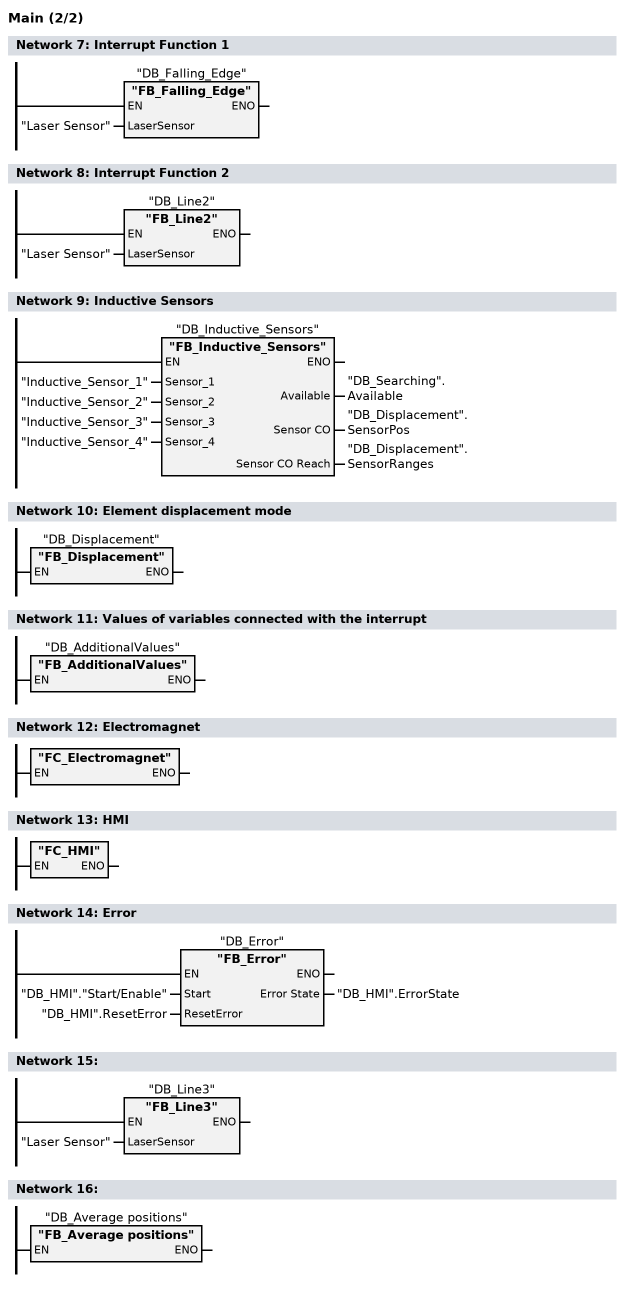
   RUNG wire#powerrail
      "DB_Falling_Edge"(LaserSensor := "Laser Sensor")
   END_RUNG
   // the same network as SCL:
   "DB_Falling_Edge"(LaserSensor := "Laser Sensor");   // "FB_Falling_Edge"
END_REGION

REGION Network 8: Interrupt Function 2
   RUNG wire#powerrail
      "DB_Line2"(LaserSensor := "Laser Sensor")
   END_RUNG
   // the same network as SCL:
   "DB_Line2"(LaserSensor := "Laser Sensor");   // "FB_Line2"
END_REGION

REGION Network 9: Inductive Sensors
   RUNG wire#powerrail
      "DB_Inductive_Sensors"(Sensor_1 := "Inductive_Sensor_1", Sensor_2 := "Inductive_Sensor_2", Sensor_3 := "Inductive_Sensor_3", Sensor_4 := "Inductive_Sensor_4", Available => "DB_Searching".Available, "Sensor CO" => "DB_Displacement".SensorPos, "Sensor CO Reach" => "DB_Displacement".SensorRanges)
   END_RUNG
   // the same network as SCL:
   "DB_Inductive_Sensors"(Sensor_1 := "Inductive_Sensor_1",   // "FB_Inductive_Sensors"
                          Sensor_2 := "Inductive_Sensor_2",
                          Sensor_3 := "Inductive_Sensor_3",
                          Sensor_4 := "Inductive_Sensor_4",
                          Available => "DB_Searching".Available,
                          "Sensor CO" => "DB_Displacement".SensorPos,
                          "Sensor CO Reach" => "DB_Displacement".SensorRanges);
END_REGION

REGION Network 10: Element displacement mode
   RUNG wire#powerrail
      "DB_Displacement"()
   END_RUNG
   // the same network as SCL:
   "DB_Displacement"();   // "FB_Displacement"
END_REGION

REGION Network 11: Values of variables connected with the interrupt
   RUNG wire#powerrail
      "DB_AdditionalValues"()
   END_RUNG
   // the same network as SCL:
   "DB_AdditionalValues"();   // "FB_AdditionalValues"
END_REGION

REGION Network 12: Electromagnet
   RUNG wire#powerrail
      "FC_Electromagnet"()
   END_RUNG
   // the same network as SCL:
   "FC_Electromagnet"();
END_REGION

REGION Network 13: HMI
   RUNG wire#powerrail
      "FC_HMI"()
   END_RUNG
   // the same network as SCL:
   "FC_HMI"();
END_REGION

REGION Network 14: Error
   RUNG wire#powerrail
      "DB_Error"(Start := "DB_HMI"."Start/Enable", ResetError := "DB_HMI".ResetError, "Error State" => "DB_HMI".ErrorState)
   END_RUNG
   // the same network as SCL:
   "DB_Error"(Start := "DB_HMI"."Start/Enable",   // "FB_Error"
              ResetError := "DB_HMI".ResetError,
              "Error State" => "DB_HMI".ErrorState);
END_REGION

REGION Network 15
   RUNG wire#powerrail
      "DB_Line3"(LaserSensor := "Laser Sensor")
   END_RUNG
   // the same network as SCL:
   "DB_Line3"(LaserSensor := "Laser Sensor");   // "FB_Line3"
END_REGION

REGION Network 16
   RUNG wire#powerrail
      "DB_Average positions"()
   END_RUNG
   // the same network as SCL:
   "DB_Average positions"();   // "FB_Average positions"
END_REGION
END_ORGANIZATION_BLOCK

ORGANIZATION_BLOCK "Hardware_IT_rising_edge"   // OB40, LAD, HWProcessInterrupt
{ S7_Optimized_Access := 'TRUE' }
VERSION : 0.1
   VAR_INPUT
      LADDR : Hw_Io;   // Hardware identifier
      USI : Word;   // User structure identifier
      IChannel : USInt;   // Interrupt channel number
      EventType : Byte;   // EventType
   END_VAR
   VAR_TEMP
      rtrig_x : Bool;
   END_VAR
BEGIN

REGION Network 1: Set when rising edge was detected
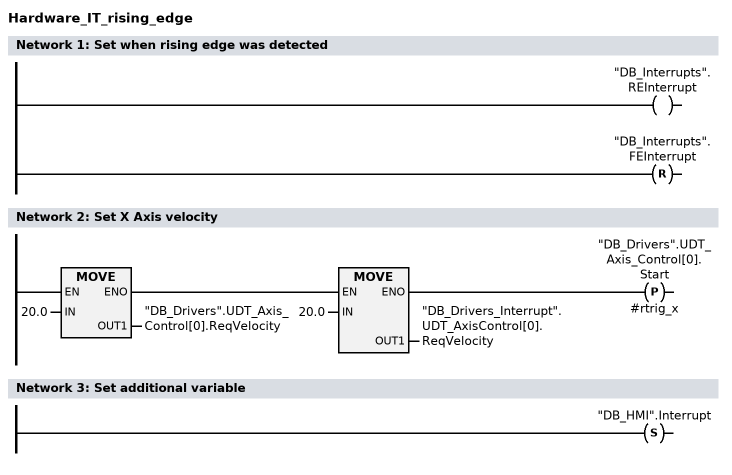
   RUNG wire#powerrail
      Coil( "DB_Interrupts".REInterrupt )
   END_RUNG
   RUNG wire#powerrail
      R_Coil( "DB_Interrupts".FEInterrupt )
   END_RUNG
   // the same network as SCL:
   "DB_Interrupts".REInterrupt := TRUE;
   "DB_Interrupts".FEInterrupt := FALSE;
END_REGION

REGION Network 2: Set X Axis velocity
   "DB_Drivers".UDT_Axis_Control[0].ReqVelocity := 20.0;
   "DB_Drivers_Interrupt".UDT_AxisControl[0].ReqVelocity := 20.0;
   "DB_Drivers".UDT_Axis_Control[0].Start := NOT #rtrig_x;   // rising edge
   #rtrig_x := TRUE;
END_REGION

REGION Network 3: Set additional variable
   RUNG wire#powerrail
      S_Coil( "DB_HMI".Interrupt )
   END_RUNG
   // the same network as SCL:
   "DB_HMI".Interrupt := TRUE;
END_REGION
END_ORGANIZATION_BLOCK

ORGANIZATION_BLOCK "Hardware_IT_falling_edge"   // OB41, LAD, HWProcessInterrupt
{ S7_Optimized_Access := 'TRUE' }
VERSION : 0.1
   VAR_INPUT
      LADDR : Hw_Io;   // Hardware identifier
      USI : Word;   // User structure identifier
      IChannel : USInt;   // Interrupt channel number
      EventType : Byte;   // EventType
   END_VAR
   VAR_TEMP
      X_Position1 : Real;
      X_Position2 : Real;
      X_Position3 : Real;
      X_Position4 : Real;
      Y_Position1 : Real;
      Y_Position2 : Real;
      Y_Position3 : Real;
      Y_Position4 : Real;
      PosReach : Bool;
      MoveX : Real;
      DelayOm : Bool;
      DelayOff : Bool;
      DebInput : Bool;
      rtrig : Bool;
      licznik : Bool;
      DontPulse : Bool;
      pulse : Bool;
      "rtrig 1" : Bool;
      diff : Real;
      i : Int;
      DontPulse2 : Bool;
      Pulse2 : Bool;
      Rtrig2 : Bool;
      j : Int;
   END_VAR
   VAR CONSTANT
      false : Bool;
      true : Bool := true;
   END_VAR
   VAR_TEMP   // added for the SCL form of the ladder/FBD networks
      _w1 : Bool;
      _w2 : Bool;
   END_VAR
BEGIN

REGION Network 1
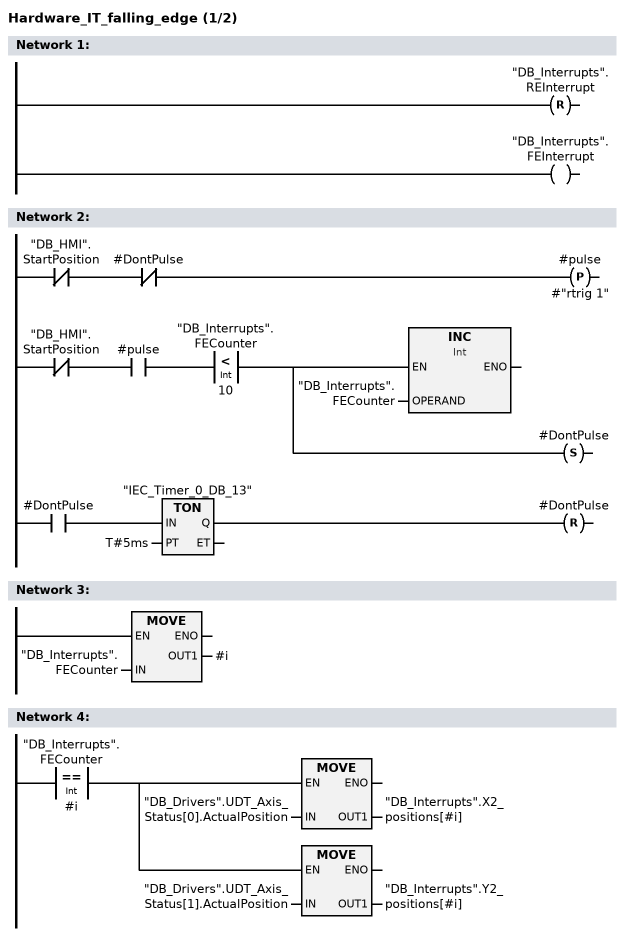
   RUNG wire#powerrail
      R_Coil( "DB_Interrupts".REInterrupt )
   END_RUNG
   RUNG wire#powerrail
      Coil( "DB_Interrupts".FEInterrupt )
   END_RUNG
   // the same network as SCL:
   "DB_Interrupts".REInterrupt := FALSE;
   "DB_Interrupts".FEInterrupt := TRUE;
END_REGION

REGION Network 2
   #_w1 := NOT "DB_HMI".StartPosition AND NOT #DontPulse;
   #pulse := #_w1 AND NOT #"rtrig 1";   // rising edge
   #"rtrig 1" := #_w1;
   #_w2 := NOT "DB_HMI".StartPosition AND #pulse AND ("DB_Interrupts".FECounter < 10);
   IF #_w2 THEN
       "DB_Interrupts".FECounter := "DB_Interrupts".FECounter + 1;
       #DontPulse := TRUE;
   END_IF;
   "IEC_Timer_0_DB_13".TON(IN := #DontPulse, PT := T#5ms);
   IF "IEC_Timer_0_DB_13".Q THEN #DontPulse := FALSE; END_IF;
END_REGION

REGION Network 3
   RUNG wire#powerrail
      Move(in := "DB_Interrupts".FECounter, out1 => #i)
   END_RUNG
   // the same network as SCL:
   #i := "DB_Interrupts".FECounter;
END_REGION

REGION Network 4
   RUNG wire#powerrail
      { S7_Templates := "SrcType := Int" } EQ_Contact(in1 := "DB_Interrupts".FECounter, in2 := #i)
      wire#w1
      Move(in := "DB_Drivers".UDT_Axis_Status[0].ActualPosition, out1 => "DB_Interrupts".X2_positions[#i])
   END_RUNG
   RUNG wire#w1
      Move(in := "DB_Drivers".UDT_Axis_Status[1].ActualPosition, out1 => "DB_Interrupts".Y2_positions[#i])
   END_RUNG
   // the same network as SCL:
   #_w1 := "DB_Interrupts".FECounter = #i;
   IF #_w1 THEN
       "DB_Interrupts".X2_positions[#i] := "DB_Drivers".UDT_Axis_Status[0].ActualPosition;
       "DB_Interrupts".Y2_positions[#i] := "DB_Drivers".UDT_Axis_Status[1].ActualPosition;
   END_IF;
END_REGION

REGION Network 5
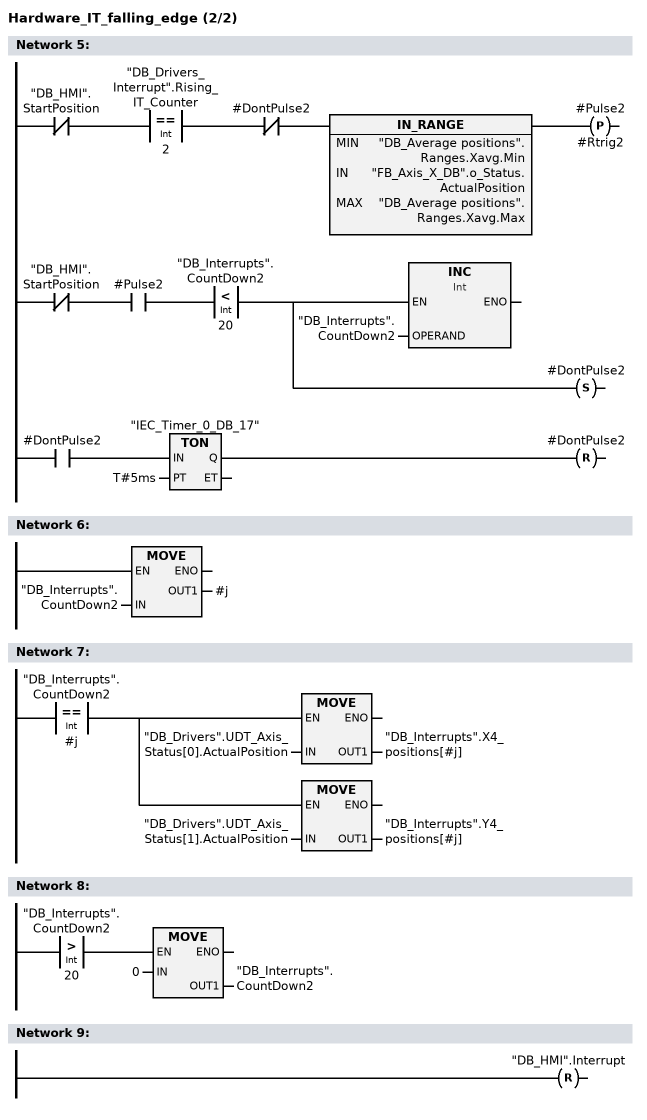
   #_w1 := NOT "DB_HMI".StartPosition AND ("DB_Drivers_Interrupt".Rising_IT_Counter = 2) AND NOT #DontPulse2 AND ("DB_Average positions".Ranges.Xavg.Min <= "FB_Axis_X_DB".o_Status.ActualPosition) AND ("FB_Axis_X_DB".o_Status.ActualPosition <= "DB_Average positions".Ranges.Xavg.Max);
   #Pulse2 := #_w1 AND NOT #Rtrig2;   // rising edge
   #Rtrig2 := #_w1;
   #_w2 := NOT "DB_HMI".StartPosition AND #Pulse2 AND ("DB_Interrupts".CountDown2 < 20);
   IF #_w2 THEN
       "DB_Interrupts".CountDown2 := "DB_Interrupts".CountDown2 + 1;
       #DontPulse2 := TRUE;
   END_IF;
   "IEC_Timer_0_DB_17".TON(IN := #DontPulse2, PT := T#5ms);
   IF "IEC_Timer_0_DB_17".Q THEN #DontPulse2 := FALSE; END_IF;
END_REGION

REGION Network 6
   RUNG wire#powerrail
      Move(in := "DB_Interrupts".CountDown2, out1 => #j)
   END_RUNG
   // the same network as SCL:
   #j := "DB_Interrupts".CountDown2;
END_REGION

REGION Network 7
   RUNG wire#powerrail
      { S7_Templates := "SrcType := Int" } EQ_Contact(in1 := "DB_Interrupts".CountDown2, in2 := #j)
      wire#w1
      Move(in := "DB_Drivers".UDT_Axis_Status[0].ActualPosition, out1 => "DB_Interrupts".X4_positions[#j])
   END_RUNG
   RUNG wire#w1
      Move(in := "DB_Drivers".UDT_Axis_Status[1].ActualPosition, out1 => "DB_Interrupts".Y4_positions[#j])
   END_RUNG
   // the same network as SCL:
   #_w1 := "DB_Interrupts".CountDown2 = #j;
   IF #_w1 THEN
       "DB_Interrupts".X4_positions[#j] := "DB_Drivers".UDT_Axis_Status[0].ActualPosition;
       "DB_Interrupts".Y4_positions[#j] := "DB_Drivers".UDT_Axis_Status[1].ActualPosition;
   END_IF;
END_REGION

REGION Network 8
   RUNG wire#powerrail
      { S7_Templates := "SrcType := Int" } GT_Contact(in1 := "DB_Interrupts".CountDown2, in2 := 20)
      Move(in := 0, out1 => "DB_Interrupts".CountDown2)
   END_RUNG
   // the same network as SCL:
   IF "DB_Interrupts".CountDown2 > 20 THEN "DB_Interrupts".CountDown2 := 0; END_IF;
END_REGION

REGION Network 9
   RUNG wire#powerrail
      R_Coil( "DB_HMI".Interrupt )
   END_RUNG
   // the same network as SCL:
   "DB_HMI".Interrupt := FALSE;
END_REGION
END_ORGANIZATION_BLOCK

// folder: RESET

FUNCTION_BLOCK "FB_RESET"   // FB6, LAD
{ S7_Optimized_Access := 'TRUE' }
VERSION : 0.1
   VAR_INPUT
      ix_StartPosition : Bool;
   END_VAR
   VAR
      Starting : Bool;
      UDT_Axis_Control : Array[0..2] of "UDT_AxisControl";
      UDT_Axis_Status : Array[0..2] of "UDT_AxisStatus";
      Rtrig : Bool;
      Start : Bool;
      Start2 : Bool;
      Rtrig2 : Bool;
      LimitY : Real;
   END_VAR
BEGIN

REGION Network 1
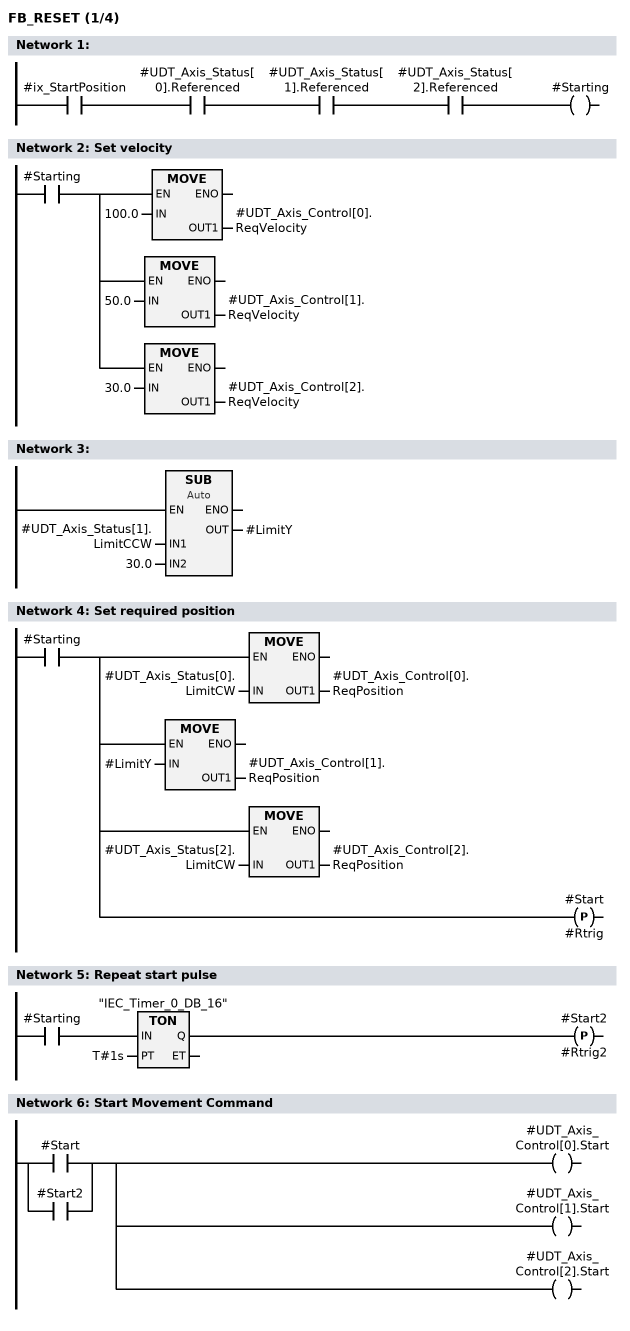
   RUNG wire#powerrail
      Contact( #ix_StartPosition )
      Contact( #UDT_Axis_Status[0].Referenced )
      Contact( #UDT_Axis_Status[1].Referenced )
      Contact( #UDT_Axis_Status[2].Referenced )
      Coil( #Starting )
   END_RUNG
   // the same network as SCL:
   #Starting := #ix_StartPosition AND #UDT_Axis_Status[0].Referenced AND #UDT_Axis_Status[1].Referenced AND #UDT_Axis_Status[2].Referenced;
END_REGION

REGION Network 2: Set velocity
   RUNG wire#powerrail
      Contact( #Starting )
      wire#w1
      Move(in := 100.0, out1 => #UDT_Axis_Control[0].ReqVelocity)
   END_RUNG
   RUNG wire#w1
      Move(in := 50.0, out1 => #UDT_Axis_Control[1].ReqVelocity)
   END_RUNG
   RUNG wire#w1
      Move(in := 30.0, out1 => #UDT_Axis_Control[2].ReqVelocity)
   END_RUNG
   // the same network as SCL:
   IF #Starting THEN
       #UDT_Axis_Control[0].ReqVelocity := 100.0;
       #UDT_Axis_Control[1].ReqVelocity := 50.0;
       #UDT_Axis_Control[2].ReqVelocity := 30.0;
   END_IF;
END_REGION

REGION Network 3
   RUNG wire#powerrail
      Sub(in1 := #UDT_Axis_Status[1].LimitCCW, in2 := 30.0, out => #LimitY)
   END_RUNG
   // the same network as SCL:
   #LimitY := #UDT_Axis_Status[1].LimitCCW - 30.0;
END_REGION

REGION Network 4: Set required position
   IF #Starting THEN
       #UDT_Axis_Control[0].ReqPosition := #UDT_Axis_Status[0].LimitCW;
       #UDT_Axis_Control[1].ReqPosition := #LimitY;
       #UDT_Axis_Control[2].ReqPosition := #UDT_Axis_Status[2].LimitCW;
   END_IF;
   #Start := #Starting AND NOT #Rtrig;   // rising edge
   #Rtrig := #Starting;
END_REGION

REGION Network 5: Repeat start pulse
   "IEC_Timer_0_DB_16".TON(IN := #Starting, PT := T#1s);
   #Start2 := "IEC_Timer_0_DB_16".Q AND NOT #Rtrig2;   // rising edge
   #Rtrig2 := "IEC_Timer_0_DB_16".Q;
END_REGION

REGION Network 6: Start Movement Command
   RUNG wire#powerrail
      Contact( #Start )
      wire#w1
      Coil( #UDT_Axis_Control[0].Start )
   END_RUNG
   RUNG wire#powerrail
      Contact( #Start2 )
   END_RUNG wire#w1
   RUNG wire#w1
      Coil( #UDT_Axis_Control[1].Start )
   END_RUNG
   RUNG wire#w1
      Coil( #UDT_Axis_Control[2].Start )
   END_RUNG
   // the same network as SCL:
   #UDT_Axis_Control[0].Start := #Start OR #Start2;
   #UDT_Axis_Control[1].Start := #Start OR #Start2;
   #UDT_Axis_Control[2].Start := #Start OR #Start2;
END_REGION

REGION Network 7: Reset variables
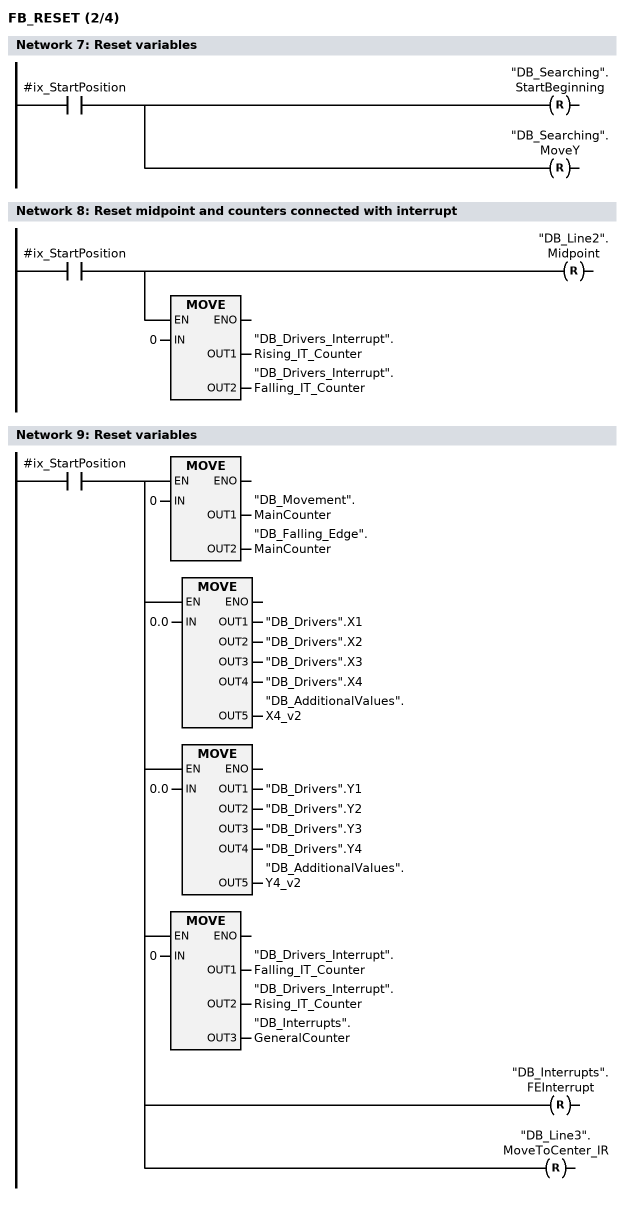
   RUNG wire#powerrail
      Contact( #ix_StartPosition )
      wire#w1
      R_Coil( "DB_Searching".StartBeginning )
   END_RUNG
   RUNG wire#w1
      R_Coil( "DB_Searching".MoveY )
   END_RUNG
   // the same network as SCL:
   IF #ix_StartPosition THEN
       "DB_Searching".StartBeginning := FALSE;
       "DB_Searching".MoveY := FALSE;
   END_IF;
END_REGION

REGION Network 8: Reset midpoint and counters connected with interrupt
   RUNG wire#powerrail
      Contact( #ix_StartPosition )
      wire#w1
      R_Coil( "DB_Line2".Midpoint )
   END_RUNG
   RUNG wire#w1
      Move(in := 0, out1 => "DB_Drivers_Interrupt".Rising_IT_Counter, out2 => "DB_Drivers_Interrupt".Falling_IT_Counter)
   END_RUNG
   // the same network as SCL:
   IF #ix_StartPosition THEN
       "DB_Line2".Midpoint := FALSE;
       "DB_Drivers_Interrupt".Rising_IT_Counter := 0;
       "DB_Drivers_Interrupt".Falling_IT_Counter := 0;
   END_IF;
END_REGION

REGION Network 9: Reset variables
   RUNG wire#powerrail
      Contact( #ix_StartPosition )
      wire#w1
      Move(in := 0, out1 => "DB_Movement".MainCounter, out2 => "DB_Falling_Edge".MainCounter)
   END_RUNG
   RUNG wire#w1
      Move(in := 0.0, out1 => "DB_Drivers".X1, out2 => "DB_Drivers".X2, out3 => "DB_Drivers".X3, out4 => "DB_Drivers".X4, out5 => "DB_AdditionalValues".X4_v2)
   END_RUNG
   RUNG wire#w1
      Move(in := 0.0, out1 => "DB_Drivers".Y1, out2 => "DB_Drivers".Y2, out3 => "DB_Drivers".Y3, out4 => "DB_Drivers".Y4, out5 => "DB_AdditionalValues".Y4_v2)
   END_RUNG
   RUNG wire#w1
      Move(in := 0, out1 => "DB_Drivers_Interrupt".Falling_IT_Counter, out2 => "DB_Drivers_Interrupt".Rising_IT_Counter, out3 => "DB_Interrupts".GeneralCounter)
   END_RUNG
   RUNG wire#w1
      R_Coil( "DB_Interrupts".FEInterrupt )
   END_RUNG
   RUNG wire#w1
      R_Coil( "DB_Line3".MoveToCenter_IR )
   END_RUNG
   // the same network as SCL:
   IF #ix_StartPosition THEN
       "DB_Movement".MainCounter := 0;
       "DB_Falling_Edge".MainCounter := 0;
       "DB_Drivers".X1 := 0.0;
       "DB_Drivers".X2 := 0.0;
       "DB_Drivers".X3 := 0.0;
       "DB_Drivers".X4 := 0.0;
       "DB_AdditionalValues".X4_v2 := 0.0;
       "DB_Drivers".Y1 := 0.0;
       "DB_Drivers".Y2 := 0.0;
       "DB_Drivers".Y3 := 0.0;
       "DB_Drivers".Y4 := 0.0;
       "DB_AdditionalValues".Y4_v2 := 0.0;
       "DB_Drivers_Interrupt".Falling_IT_Counter := 0;
       "DB_Drivers_Interrupt".Rising_IT_Counter := 0;
       "DB_Interrupts".GeneralCounter := 0;
       "DB_Interrupts".FEInterrupt := FALSE;
       "DB_Line3".MoveToCenter_IR := FALSE;
   END_IF;
END_REGION

REGION Network 10: Reset remembered occupied place if reset button was pressed
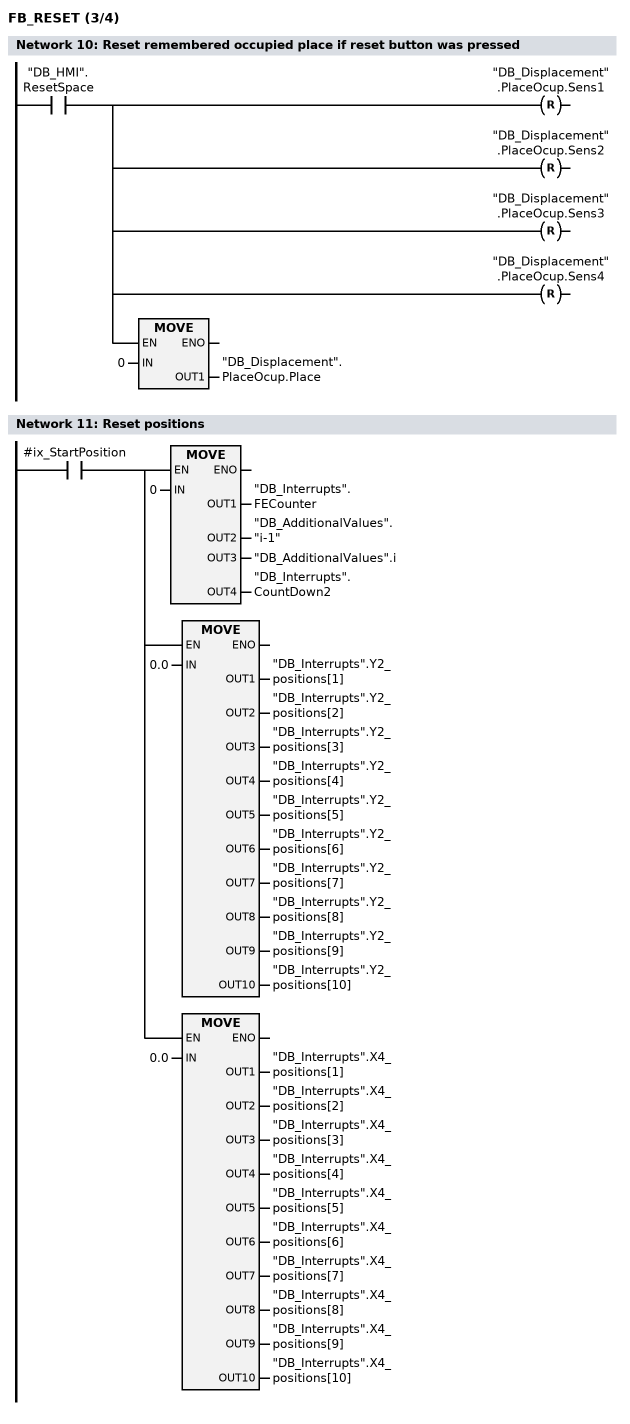
   RUNG wire#powerrail
      Contact( "DB_HMI".ResetSpace )
      wire#w1
      R_Coil( "DB_Displacement".PlaceOcup.Sens1 )
   END_RUNG
   RUNG wire#w1
      R_Coil( "DB_Displacement".PlaceOcup.Sens2 )
   END_RUNG
   RUNG wire#w1
      R_Coil( "DB_Displacement".PlaceOcup.Sens3 )
   END_RUNG
   RUNG wire#w1
      R_Coil( "DB_Displacement".PlaceOcup.Sens4 )
   END_RUNG
   RUNG wire#w1
      Move(in := 0, out1 => "DB_Displacement".PlaceOcup.Place)
   END_RUNG
   // the same network as SCL:
   IF "DB_HMI".ResetSpace THEN
       "DB_Displacement".PlaceOcup.Sens1 := FALSE;
       "DB_Displacement".PlaceOcup.Sens2 := FALSE;
       "DB_Displacement".PlaceOcup.Sens3 := FALSE;
       "DB_Displacement".PlaceOcup.Sens4 := FALSE;
       "DB_Displacement".PlaceOcup.Place := 0;
   END_IF;
END_REGION

REGION Network 11: Reset positions
   RUNG wire#powerrail
      Contact( #ix_StartPosition )
      wire#w1
      Move(in := 0, out1 => "DB_Interrupts".FECounter, out2 => "DB_AdditionalValues"."i-1", out3 => "DB_AdditionalValues".i, out4 => "DB_Interrupts".CountDown2)
   END_RUNG
   RUNG wire#w1
      Move(in := 0.0, out1 => "DB_Interrupts".Y2_positions[1], out2 => "DB_Interrupts".Y2_positions[2], out3 => "DB_Interrupts".Y2_positions[3], out4 => "DB_Interrupts".Y2_positions[4], out5 => "DB_Interrupts".Y2_positions[5], out6 => "DB_Interrupts".Y2_positions[6], out7 => "DB_Interrupts".Y2_positions[7], out8 => "DB_Interrupts".Y2_positions[8], out9 => "DB_Interrupts".Y2_positions[9], out10 => "DB_Interrupts".Y2_positions[10])
   END_RUNG
   RUNG wire#w1
      Move(in := 0.0, out1 => "DB_Interrupts".X4_positions[1], out2 => "DB_Interrupts".X4_positions[2], out3 => "DB_Interrupts".X4_positions[3], out4 => "DB_Interrupts".X4_positions[4], out5 => "DB_Interrupts".X4_positions[5], out6 => "DB_Interrupts".X4_positions[6], out7 => "DB_Interrupts".X4_positions[7], out8 => "DB_Interrupts".X4_positions[8], out9 => "DB_Interrupts".X4_positions[9], out10 => "DB_Interrupts".X4_positions[10])
   END_RUNG
   // the same network as SCL:
   IF #ix_StartPosition THEN
       "DB_Interrupts".FECounter := 0;
       "DB_AdditionalValues"."i-1" := 0;
       "DB_AdditionalValues".i := 0;
       "DB_Interrupts".CountDown2 := 0;
       "DB_Interrupts".Y2_positions[1] := 0.0;
       "DB_Interrupts".Y2_positions[2] := 0.0;
       "DB_Interrupts".Y2_positions[3] := 0.0;
       "DB_Interrupts".Y2_positions[4] := 0.0;
       "DB_Interrupts".Y2_positions[5] := 0.0;
       "DB_Interrupts".Y2_positions[6] := 0.0;
       "DB_Interrupts".Y2_positions[7] := 0.0;
       "DB_Interrupts".Y2_positions[8] := 0.0;
       "DB_Interrupts".Y2_positions[9] := 0.0;
       "DB_Interrupts".Y2_positions[10] := 0.0;
       "DB_Interrupts".X4_positions[1] := 0.0;
       "DB_Interrupts".X4_positions[2] := 0.0;
       "DB_Interrupts".X4_positions[3] := 0.0;
       "DB_Interrupts".X4_positions[4] := 0.0;
       "DB_Interrupts".X4_positions[5] := 0.0;
       "DB_Interrupts".X4_positions[6] := 0.0;
       "DB_Interrupts".X4_positions[7] := 0.0;
       "DB_Interrupts".X4_positions[8] := 0.0;
       "DB_Interrupts".X4_positions[9] := 0.0;
       "DB_Interrupts".X4_positions[10] := 0.0;
   END_IF;
END_REGION

REGION Network 12: Reset variables
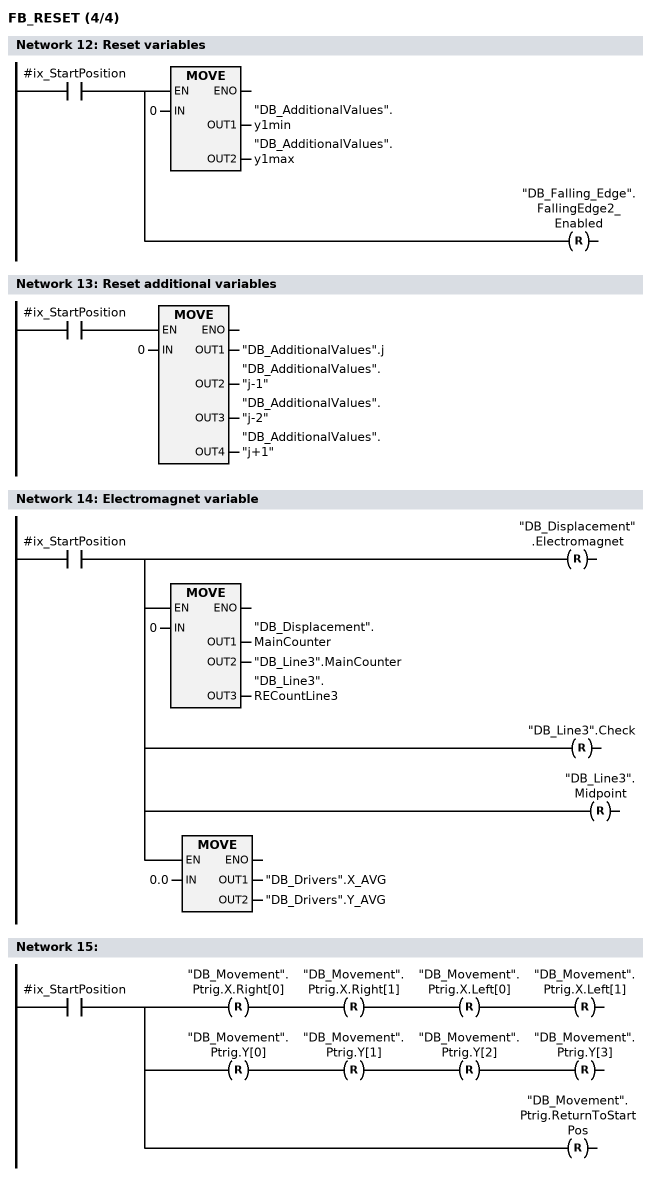
   RUNG wire#powerrail
      Contact( #ix_StartPosition )
      wire#w1
      Move(in := 0, out1 => "DB_AdditionalValues".y1min, out2 => "DB_AdditionalValues".y1max)
   END_RUNG
   RUNG wire#w1
      R_Coil( "DB_Falling_Edge".FallingEdge2_Enabled )
   END_RUNG
   // the same network as SCL:
   IF #ix_StartPosition THEN
       "DB_AdditionalValues".y1min := 0;
       "DB_AdditionalValues".y1max := 0;
       "DB_Falling_Edge".FallingEdge2_Enabled := FALSE;
   END_IF;
END_REGION

REGION Network 13: Reset additional variables
   RUNG wire#powerrail
      Contact( #ix_StartPosition )
      Move(in := 0, out1 => "DB_AdditionalValues".j, out2 => "DB_AdditionalValues"."j-1", out3 => "DB_AdditionalValues"."j-2", out4 => "DB_AdditionalValues"."j+1")
   END_RUNG
   // the same network as SCL:
   IF #ix_StartPosition THEN
       "DB_AdditionalValues".j := 0;
       "DB_AdditionalValues"."j-1" := 0;
       "DB_AdditionalValues"."j-2" := 0;
       "DB_AdditionalValues"."j+1" := 0;
   END_IF;
END_REGION

REGION Network 14: Electromagnet variable
   RUNG wire#powerrail
      Contact( #ix_StartPosition )
      wire#w1
      R_Coil( "DB_Displacement".Electromagnet )
   END_RUNG
   RUNG wire#w1
      Move(in := 0, out1 => "DB_Displacement".MainCounter, out2 => "DB_Line3".MainCounter, out3 => "DB_Line3".RECountLine3)
   END_RUNG
   RUNG wire#w1
      R_Coil( "DB_Line3".Check )
   END_RUNG
   RUNG wire#w1
      R_Coil( "DB_Line3".Midpoint )
   END_RUNG
   RUNG wire#w1
      Move(in := 0.0, out1 => "DB_Drivers".X_AVG, out2 => "DB_Drivers".Y_AVG)
   END_RUNG
   // the same network as SCL:
   IF #ix_StartPosition THEN
       "DB_Displacement".Electromagnet := FALSE;
       "DB_Displacement".MainCounter := 0;
       "DB_Line3".MainCounter := 0;
       "DB_Line3".RECountLine3 := 0;
       "DB_Line3".Check := FALSE;
       "DB_Line3".Midpoint := FALSE;
       "DB_Drivers".X_AVG := 0.0;
       "DB_Drivers".Y_AVG := 0.0;
   END_IF;
END_REGION

REGION Network 15
   RUNG wire#powerrail
      Contact( #ix_StartPosition )
      wire#w1
      R_Coil( "DB_Movement".Ptrig.X.Right[0] )
      R_Coil( "DB_Movement".Ptrig.X.Right[1] )
      R_Coil( "DB_Movement".Ptrig.X.Left[0] )
      R_Coil( "DB_Movement".Ptrig.X.Left[1] )
   END_RUNG
   RUNG wire#w1
      R_Coil( "DB_Movement".Ptrig.Y[0] )
      R_Coil( "DB_Movement".Ptrig.Y[1] )
      R_Coil( "DB_Movement".Ptrig.Y[2] )
      R_Coil( "DB_Movement".Ptrig.Y[3] )
   END_RUNG
   RUNG wire#w1
      R_Coil( "DB_Movement".Ptrig.ReturnToStartPos )
   END_RUNG
   // the same network as SCL:
   IF #ix_StartPosition THEN
       "DB_Movement".Ptrig.X.Right[0] := FALSE;
       "DB_Movement".Ptrig.X.Right[1] := FALSE;
       "DB_Movement".Ptrig.X.Left[0] := FALSE;
       "DB_Movement".Ptrig.X.Left[1] := FALSE;
       "DB_Movement".Ptrig.Y[0] := FALSE;
       "DB_Movement".Ptrig.Y[1] := FALSE;
       "DB_Movement".Ptrig.Y[2] := FALSE;
       "DB_Movement".Ptrig.Y[3] := FALSE;
       "DB_Movement".Ptrig.ReturnToStartPos := FALSE;
   END_IF;
END_REGION
END_FUNCTION_BLOCK

// folder: Searching Mode

FUNCTION_BLOCK "FB_Searching"   // FB2, LAD
{ S7_Optimized_Access := 'TRUE' }